DATA_BLOCK "Recipe Libraries"   // DB9
{ S7_Optimized_Access := 'TRUE' }
VERSION : 0.1
   VAR
      me : "Menu: Libraries";
   END_VAR
BEGIN
   me.stations[24].wip[0] := WSTRING#'16.08.208.101.020A$L$$SA DOC Sleeved Before Forming';
   me.stations[24].wip[1] := WSTRING#'16.08.209.031.000C$LDOC Stuffed Shell Before Forming';
   me.stations[24].wip[2] := WSTRING#'16.08.209.091.000D$LSA DPF Stuffed (after Hess)';
   me.stations[24].wip[3] := WSTRING#'16.08.209.233.000E$LSCR Stuffed Shell- NGK Before Forming';
   me.stations[24].wip[4] := WSTRING#'16.08.209.437.000A$LDOC Stuffed Shell Unformed';
   me.stations[24].wip[5] := WSTRING#'16.08.210.031.000B$LStuffed Shell DOC';
   me.stations[24].wip[6] := WSTRING#'16.08.210.421.500A$LStuffed Shell DOC- 2013';
   me.stations[24].wip[7] := WSTRING#'16.08.210.428.000A$LSA DPF Stuffed (after Hess)';
   me.stations[24].wip[8] := WSTRING#'16.08.211.801.400A$L$$SA DOC Sleeved';
   me.stations[24].wip[9] := WSTRING#'16.08.211.801.700B$LDPF Stuffed Shell 1 box longs only';
   me.stations[24].wip[10] := WSTRING#'16.08.211.806.400B$L$$SA DPF Stuffed Shell';
   me.stations[24].wip[11] := WSTRING#'16.08.216.801.600A$LSA DOC Sleeved DDC 2016 unformed';
   me.stations[24].wip[12] := WSTRING#'16.08.216.806.400A$L DPF Sleeved 2016';
   me.stations[24].wip[13] := WSTRING#'16.08.217.408.000A$LSA DPF SLEEVED Hess';
   me.stations[24].wip[14] := WSTRING#'16.08.217.421.500A$LSA DOC SLEEVED - 2HH 2016';
   me.stations[24].wip[15] := WSTRING#'16.08.217.737.000A$LSA DOC SLEEVED - 2V2 2016 unformed';
   me.stations[24].wip[16] := WSTRING#'16.32.307.322.210A$LVolvo - ASSY INLET - SUB 8 Unformed';
   me.stations[24].wip[17] := WSTRING#'16.32.307.332.400A$LAssembly DPF Canning 2016';
   me.stations[24].wip[18] := WSTRING#'16.32.307.472.210A$LSA DOC Canning w/out End Forming';
   me.stations[24].wip[19] := WSTRING#'16.32.407.322.210A$LVOLVO DOC STUFFED SHELL UNFORMED';
   me.stations[24].wip[20] := WSTRING#'16.08.208.081.000H$LDPF Stuffed Shell 1 box longs only';
   me.stations[24].wip[21] := WSTRING#'16.08.208.621.000G$LSA DPF Stuffed Shell';
   me.stations[24].wip[22] := WSTRING#'16.32.407.322.300A$LDPF Stuffed Shell: MD13/MD16';
   me.stations[24].wip[23] := WSTRING#'16.32.307.332.300A$LDPF Stuffed Shell MD11';
   me.stations[25].wip[0] := WSTRING#'16.08.210.421.500A$LStuffed Shell DOC- 2013';
   me.stations[25].wip[1] := WSTRING#'16.08.217.421.500A$LSA DOC SLEEVED - 2HH 2016';
   me.stations[25].wip[2] := WSTRING#'16.08.217.737.000A$LSA DOC SLEEVED - 2V2 2016 unformed';
   me.stations[25].wip[3] := WSTRING#'16.08.208.031.000F$LSCR Stuffed Shell 1 box longs only';
   me.stations[25].wip[4] := WSTRING#'16.08.208.651.000G$LStuffed Shell SCR- NGK';
   me.stations[25].wip[5] := WSTRING#'16.08.211.803.400A$LSCR Stuffed Shell High Power';
   me.stations[25].wip[6] := WSTRING#'16.08.217.233.000A$LSA SCR SLEEVED before FORMING';
   me.stations[25].wip[7] := WSTRING#'16.32.606.411.000A$LStuffed Shell - SCR Horizontal';
   me.stations[25].wip[8] := WSTRING#'16.32.606.421.000A$LStuffed Shell - SCR Horizontal Long- UNI';
   me.stations[25].wip[9] := WSTRING#'16.32.706.311.000A$L$$SCR Stuffed Shell MD11/13: Vert Short';
   me.stations[25].wip[10] := WSTRING#'16.32.706.311.001A$L$$SCR Stuffed Shell MD11/13: Vert Short';
   me.stations[25].wip[11] := WSTRING#'16.32.706.341.000A$LSA SCR Catalyst Module - MD11_MD13 -';
   me.stations[25].wip[12] := WSTRING#'16.32.706.401.000A$LSCR Stuffed Shell MD11/13: Australia';
   me.stations[26].wip[0] := WSTRING#'16.18.015.420.000A$LSA DOC CANNING 11.25 x 5in -END FORMED-';
   me.stations[26].wip[1] := WSTRING#'16.08.211.806.400B$L$$SA DPF Stuffed Shell';
   me.stations[26].wip[2] := WSTRING#'16.08.216.801.600A$LSA DOC Sleeved DDC 2016 unformed';
   me.stations[26].wip[3] := WSTRING#'16.08.216.806.400A$L DPF Sleeved 2016';
   me.stations[26].wip[4] := WSTRING#'16.08.216.751.100A$LSA Sleeved SCR 2016';
   me.stations[26].wip[5] := WSTRING#'16.18.007.300.000A$LSA SCR CANNING 9.5 x 10in -END FORMED-';
   me.stations[26].wip[6] := WSTRING#'16.18.007.310.000A$LSA SCR CANNING 9.5 x 12in -END FORMED-';
   me.stations[26].wip[7] := WSTRING#'16.18.007.320.000B$LSA SCR CANNING 9.5 x 9in -END FORMED-';
   me.stations[26].wip[8] := WSTRING#'16.18.008.300.000A$LSA SCR CANNING 9.5 x 12in -END FORMED-';
   me.stations[26].wip[9] := WSTRING#'16.18.008.310.000A$LSA SCR CANNING 9.5 x 10in -END FORMED-';
   me.stations[26].wip[10] := WSTRING#'16.18.008.320.000A$LSA SCR CANNING 9.5 x 13in -END FORMED-';
   me.stations[26].wip[11] := WSTRING#'16.18.008.340.000A$LSA SCR CANNING 9.5 x 13in -END FORMED-';
   me.stations[26].wip[12] := WSTRING#'16.18.009.301.000H$LSA SCR CANNING 13 x 11in UNFORMED-';
   me.stations[26].wip[13] := WSTRING#'16.18.009.311.000H$LSA SCR CANNING 13 x 12in UNFORMED-';
   me.stations[26].wip[14] := WSTRING#'16.18.009.321.000G$LSA SCR CANNING 13 x 9in UNFORMED';
   me.stations[26].wip[15] := WSTRING#'16.18.009.331.000F$LSA SCR CANNING 13 x 9in UNFORMED';
   me.stations[26].wip[16] := WSTRING#'16.18.009.371.000D$LSA SCR CANNING 13 X10  UNFORMED';
   me.stations[26].wip[17] := WSTRING#'16.18.011.300.000A$LSA SCR CANNING 9.5 x 13.5in -END FORMED-';
   me.stations[26].wip[18] := WSTRING#'16.18.011.310.000A$L SA SCR CANNING 9.5 x 10in -END FORMED-';
   me.stations[26].wip[19] := WSTRING#'16.18.011.320.000A$LSA SCR CANNING 9_5 x 13in -END FORMED-';
   me.stations[26].wip[20] := WSTRING#'16.18.011.330.000A$LSA SCR CANNING 9.5 x 9in -END FORMED-';
   me.stations[26].wip[21] := WSTRING#'16.18.012.400.000A$LSA DOC CANNING 9.5 x 4in -END FORMED_';
   me.stations[26].wip[22] := WSTRING#'16.18.012.410.000A$LSA DOC CANNING 9.5 x 3.3in -END FORMED-';
   me.stations[26].wip[23] := WSTRING#'16.18.012.420.000A$LSA DOC CANNING 9.5 x 4in -END FORMED-';
   me.stations[26].wip[24] := WSTRING#'16.18.012.430.000A$LSA DOC CANNING 9.5 x 3.3in -END FORMED-';
   me.stations[26].wip[25] := WSTRING#'16.18.012.440.000A$LSA DOC CANNING 9.5 x 5in -END FORMED-';
   me.stations[26].wip[26] := WSTRING#'16.18.013.410.000A$LSA DOC CANNING 9_5 x 4_5in -END FORMED-';
   me.stations[26].wip[27] := WSTRING#'16.18.013.420.000A$LSA DOC CANNING 9.5 x 5.5in -END FORMED-';
   me.stations[26].wip[28] := WSTRING#'16.18.015.400.000A$LSA DOC CANNING 11.25 x 4in -END FORMED-';
   me.stations[26].wip[29] := WSTRING#'16.18.015.410.000A$LSA DOC CANNING 11_25 x 5in -END FORMED-';
   me.stations[26].wip[30] := WSTRING#'16.18.015.430.000A$LSA DOC CANNING 11.25 x 3.4in -END FORMED';
   me.stations[26].wip[31] := WSTRING#'16.18.015.450.000A$LSA DOC CANNING 11.25 x 5in -END FORMED-';
   me.stations[26].wip[32] := WSTRING#'16.18.016.400.000A$LSA DOC CANNING 11.25 x 3.4in -END FORMED';
   me.stations[26].wip[33] := WSTRING#'16.18.017.300.000A$LSA SCR CANNING 12 x 10in -END FORMED-';
   me.stations[26].wip[34] := WSTRING#'16.18.017.310.000A$LSA SCR CANNING 12 x 9in -END FORMED-';
   me.stations[26].wip[35] := WSTRING#'16.18.017.321.000F$LSA SCR CANNING 12x7in UNFORMED-';
   me.stations[26].wip[36] := WSTRING#'16.18.018.400.000A$LSA DOC CANNING 11.25 x 6.8in -END FORMED';
   me.stations[26].wip[37] := WSTRING#'16.18.018.410.000A$LSA DOC CANNING 11.25 x 5in -END FORMED-';
   me.stations[26].wip[38] := WSTRING#'16.18.018.420.000A$LSA DOC CANNING 11.25 x 6.8in -END FORMED';
   me.stations[26].wip[39] := WSTRING#'16.18.018.440.000A$LSA DOC CANNING 11.25 x 5in -END FORMED-';
   me.stations[26].wip[40] := WSTRING#'16.18.011.340.000A$LSCR CANNING 9.5 x 9in -END FORMED-';
   me.stations[27].wip[0] := WSTRING#'16.08.211.801.700B$LDPF Stuffed Shell 1 box longs only';
   me.stations[27].wip[1] := WSTRING#'16.32.307.322.210A$LVolvo - ASSY INLET - SUB 8 Unformed';
   me.stations[27].wip[2] := WSTRING#'16.32.606.411.000A$LStuffed Shell - SCR Horizontal';
   me.stations[27].wip[3] := WSTRING#'16.32.112.311.001A$LSA SCR CANNING UNFORMED';
   me.stations[27].wip[4] := WSTRING#'16.32.112.553.300C$LSA SCR CANNING A700 UNFORMED';
   me.stations[27].wip[5] := WSTRING#'16.32.112.304.008A$LASSY SCR CANNING FORMED';
   me.stations[27].wip[6] := WSTRING#'16.32.112.516.000G$LASSY DPF CANNING A700';
   me.stations[27].wip[7] := WSTRING#'16.32.112.543.000E$LASSY DOC CANNING A700';
   me.stations[28].wip[0] := WSTRING#'11.52.001.312.000B$LSA JL 2.2L DPF CANNING';
   me.stations[28].wip[1] := WSTRING#'11.54.007.309.000D$LSTUFFED SHELL ASSEMBLY USA-U625';
   me.stations[28].wip[2] := WSTRING#'11.54.007.309.002D$LSTUFFED SHELL ASSEMBLY USA-U625';
   me.stations[28].wip[3] := WSTRING#'11.54.007.309.009D$LSTUFFED SHELL ASSEMBLY USA-U625';
   me.stations[24].raw[20,7] := WSTRING#'';
   me.stations[24].raw[20,6] := WSTRING#'';
   me.stations[24].raw[20,5] := WSTRING#'';
   me.stations[24].raw[20,4] := WSTRING#'';
   me.stations[24].raw[20,3] := WSTRING#'';
   me.stations[24].raw[20,2] := WSTRING#'16.08.208.091.000A';
   me.stations[24].raw[20,1] := WSTRING#'16.08.208.311.000F';
   me.stations[24].raw[20,0] := WSTRING#'16.08.208.081.010B';
   me.stations[24].raw[19,7] := WSTRING#'';
   me.stations[24].raw[19,6] := WSTRING#'';
   me.stations[24].raw[19,5] := WSTRING#'';
   me.stations[24].raw[19,4] := WSTRING#'';
   me.stations[24].raw[19,3] := WSTRING#'';
   me.stations[24].raw[19,2] := WSTRING#'16.32.407.241.150B';
   me.stations[24].raw[19,1] := WSTRING#'16.32.407.241.170B';
   me.stations[24].raw[19,0] := WSTRING#'16.32.407.441.160A';
   me.stations[24].raw[18,7] := WSTRING#'';
   me.stations[24].raw[18,6] := WSTRING#'';
   me.stations[24].raw[18,5] := WSTRING#'';
   me.stations[24].raw[18,4] := WSTRING#'';
   me.stations[24].raw[18,3] := WSTRING#'';
   me.stations[24].raw[18,2] := WSTRING#'16.32.112.543.020A';
   me.stations[24].raw[18,1] := WSTRING#'16.32.307.211.170B';
   me.stations[24].raw[18,0] := WSTRING#'16.32.307.461.160A';
   me.stations[24].raw[17,7] := WSTRING#'';
   me.stations[24].raw[17,6] := WSTRING#'';
   me.stations[24].raw[17,5] := WSTRING#'';
   me.stations[24].raw[17,4] := WSTRING#'';
   me.stations[24].raw[17,3] := WSTRING#'';
   me.stations[24].raw[17,2] := WSTRING#'16.32.112.536.010A';
   me.stations[24].raw[17,1] := WSTRING#'16.32.307.212.320C';
   me.stations[24].raw[17,0] := WSTRING#'16.32.307.312.310A';
   me.stations[24].raw[16,7] := WSTRING#'';
   me.stations[24].raw[16,6] := WSTRING#'';
   me.stations[24].raw[16,5] := WSTRING#'';
   me.stations[24].raw[16,4] := WSTRING#'';
   me.stations[24].raw[16,3] := WSTRING#'';
   me.stations[24].raw[16,2] := WSTRING#'16.32.307.211.150B';
   me.stations[24].raw[16,1] := WSTRING#'16.32.307.211.170B';
   me.stations[24].raw[16,0] := WSTRING#'16.32.307.461.160A';
   me.stations[24].raw[15,7] := WSTRING#'';
   me.stations[24].raw[15,6] := WSTRING#'';
   me.stations[24].raw[15,5] := WSTRING#'';
   me.stations[24].raw[15,4] := WSTRING#'';
   me.stations[24].raw[15,3] := WSTRING#'';
   me.stations[24].raw[15,2] := WSTRING#'16.08.217.421.130A';
   me.stations[24].raw[15,1] := WSTRING#'16.08.209.031.010C';
   me.stations[24].raw[15,0] := WSTRING#'16.08.209.031.030B';
   me.stations[24].raw[14,7] := WSTRING#'';
   me.stations[24].raw[14,6] := WSTRING#'';
   me.stations[24].raw[14,5] := WSTRING#'';
   me.stations[24].raw[14,4] := WSTRING#'';
   me.stations[24].raw[14,3] := WSTRING#'';
   me.stations[24].raw[14,2] := WSTRING#'16.08.217.421.130A';
   me.stations[24].raw[14,1] := WSTRING#'16.08.210.031.010B';
   me.stations[24].raw[14,0] := WSTRING#'16.08.209.031.030B';
   me.stations[24].raw[13,7] := WSTRING#'';
   me.stations[24].raw[13,6] := WSTRING#'';
   me.stations[24].raw[13,5] := WSTRING#'';
   me.stations[24].raw[13,4] := WSTRING#'';
   me.stations[24].raw[13,3] := WSTRING#'';
   me.stations[24].raw[13,2] := WSTRING#'16.08.217.421.010A';
   me.stations[24].raw[13,1] := WSTRING#'16.08.209.091.010C';
   me.stations[24].raw[13,0] := WSTRING#'16.08.210.421.020A';
   me.stations[24].raw[12,7] := WSTRING#'';
   me.stations[24].raw[12,6] := WSTRING#'';
   me.stations[24].raw[12,5] := WSTRING#'';
   me.stations[24].raw[12,4] := WSTRING#'';
   me.stations[24].raw[12,3] := WSTRING#'';
   me.stations[24].raw[12,2] := WSTRING#'16.08.216.806.020A';
   me.stations[24].raw[12,1] := WSTRING#'16.08.208.631.000F';
   me.stations[24].raw[12,0] := WSTRING#'16.08.216.315.000A';
   me.stations[24].raw[11,7] := WSTRING#'';
   me.stations[24].raw[11,6] := WSTRING#'';
   me.stations[24].raw[11,5] := WSTRING#'';
   me.stations[24].raw[11,4] := WSTRING#'';
   me.stations[24].raw[11,3] := WSTRING#'';
   me.stations[24].raw[11,2] := WSTRING#'16.08.216.053.000A';
   me.stations[24].raw[11,1] := WSTRING#'16.08.208.321.000G';
   me.stations[24].raw[11,0] := WSTRING#'16.08.208.101.010C';
   me.stations[24].raw[10,7] := WSTRING#'';
   me.stations[24].raw[10,6] := WSTRING#'';
   me.stations[24].raw[10,5] := WSTRING#'';
   me.stations[24].raw[10,4] := WSTRING#'';
   me.stations[24].raw[10,3] := WSTRING#'';
   me.stations[24].raw[10,2] := WSTRING#'16.08.211.806.020A';
   me.stations[24].raw[10,1] := WSTRING#'16.08.208.631.000F';
   me.stations[24].raw[10,0] := WSTRING#'16.08.216.315.000A';
   me.stations[24].raw[9,7] := WSTRING#'';
   me.stations[24].raw[9,6] := WSTRING#'';
   me.stations[24].raw[9,5] := WSTRING#'';
   me.stations[24].raw[9,4] := WSTRING#'';
   me.stations[24].raw[9,3] := WSTRING#'';
   me.stations[24].raw[9,2] := WSTRING#'16.08.211.801.020A';
   me.stations[24].raw[9,1] := WSTRING#'16.08.208.631.000F';
   me.stations[24].raw[9,0] := WSTRING#'16.08.216.315.002A';
   me.stations[24].raw[8,7] := WSTRING#'';
   me.stations[24].raw[8,6] := WSTRING#'';
   me.stations[24].raw[8,5] := WSTRING#'';
   me.stations[24].raw[8,4] := WSTRING#'';
   me.stations[24].raw[8,3] := WSTRING#'';
   me.stations[24].raw[8,2] := WSTRING#'16.08.211.801.010A';
   me.stations[24].raw[8,1] := WSTRING#'16.08.208.321.000G';
   me.stations[24].raw[8,0] := WSTRING#'16.08.208.101.010C';
   me.stations[24].raw[7,7] := WSTRING#'';
   me.stations[24].raw[7,6] := WSTRING#'';
   me.stations[24].raw[7,5] := WSTRING#'';
   me.stations[24].raw[7,4] := WSTRING#'';
   me.stations[24].raw[7,3] := WSTRING#'';
   me.stations[24].raw[7,2] := WSTRING#'16.08.210.421.010A';
   me.stations[24].raw[7,1] := WSTRING#'16.08.209.091.010C';
   me.stations[24].raw[7,0] := WSTRING#'16.08.210.421.020A';
   me.stations[24].raw[6,7] := WSTRING#'';
   me.stations[24].raw[6,6] := WSTRING#'';
   me.stations[24].raw[6,5] := WSTRING#'';
   me.stations[24].raw[6,4] := WSTRING#'';
   me.stations[24].raw[6,3] := WSTRING#'';
   me.stations[24].raw[6,2] := WSTRING#'16.08.210.421.030A';
   me.stations[24].raw[6,1] := WSTRING#'16.08.210.031.010B';
   me.stations[24].raw[6,0] := WSTRING#'16.08.209.031.030B';
   me.stations[24].raw[5,7] := WSTRING#'';
   me.stations[24].raw[5,6] := WSTRING#'';
   me.stations[24].raw[5,5] := WSTRING#'';
   me.stations[24].raw[5,4] := WSTRING#'';
   me.stations[24].raw[5,3] := WSTRING#'';
   me.stations[24].raw[5,2] := WSTRING#'16.08.209.031.050A';
   me.stations[24].raw[5,1] := WSTRING#'16.08.210.031.010B';
   me.stations[24].raw[5,0] := WSTRING#'16.08.209.031.030B';
   me.stations[24].raw[4,7] := WSTRING#'';
   me.stations[24].raw[4,6] := WSTRING#'';
   me.stations[24].raw[4,5] := WSTRING#'';
   me.stations[24].raw[4,4] := WSTRING#'';
   me.stations[24].raw[4,3] := WSTRING#'';
   me.stations[24].raw[4,2] := WSTRING#'16.08.210.421.030A';
   me.stations[24].raw[4,1] := WSTRING#'16.08.209.031.010C';
   me.stations[24].raw[4,0] := WSTRING#'16.08.209.031.030B';
   me.stations[24].raw[3,7] := WSTRING#'';
   me.stations[24].raw[3,6] := WSTRING#'';
   me.stations[24].raw[3,5] := WSTRING#'';
   me.stations[24].raw[3,4] := WSTRING#'16.08.208.041.000A';
   me.stations[24].raw[3,3] := WSTRING#'16.08.211.291.000A';
   me.stations[24].raw[3,2] := WSTRING#'16.08.209.232.010C';
   me.stations[24].raw[3,1] := WSTRING#'16.08.208.031.020C';
   me.stations[24].raw[3,0] := WSTRING#'16.08.208.651.010B';
   me.stations[24].raw[2,7] := WSTRING#'';
   me.stations[24].raw[2,6] := WSTRING#'';
   me.stations[24].raw[2,5] := WSTRING#'';
   me.stations[24].raw[2,4] := WSTRING#'';
   me.stations[24].raw[2,3] := WSTRING#'';
   me.stations[24].raw[2,2] := WSTRING#'16.08.209.091.060A';
   me.stations[24].raw[2,1] := WSTRING#'16.08.209.091.010C';
   me.stations[24].raw[2,0] := WSTRING#'16.08.209.091.030D';
   me.stations[24].raw[1,7] := WSTRING#'';
   me.stations[24].raw[1,6] := WSTRING#'';
   me.stations[24].raw[1,5] := WSTRING#'';
   me.stations[24].raw[1,4] := WSTRING#'';
   me.stations[24].raw[1,3] := WSTRING#'';
   me.stations[24].raw[1,2] := WSTRING#'16.08.209.031.050A';
   me.stations[24].raw[1,1] := WSTRING#'16.08.209.031.010C';
   me.stations[24].raw[1,0] := WSTRING#'16.08.209.031.030B';
   me.stations[24].raw[0,7] := WSTRING#'';
   me.stations[24].raw[0,6] := WSTRING#'';
   me.stations[24].raw[0,5] := WSTRING#'';
   me.stations[24].raw[0,4] := WSTRING#'';
   me.stations[24].raw[0,3] := WSTRING#'';
   me.stations[24].raw[0,2] := WSTRING#'16.08.208.111.000B';
   me.stations[24].raw[0,1] := WSTRING#'16.08.208.321.000G';
   me.stations[24].raw[0,0] := WSTRING#'16.08.208.101.010C';
   me.stations[26].raw[15,6] := WSTRING#'';
   me.stations[26].raw[15,5] := WSTRING#'';
   me.stations[26].raw[15,4] := WSTRING#'16.18.009.331.050A';
   me.stations[26].raw[15,3] := WSTRING#'16.18.009.321.030A';
   me.stations[26].raw[15,2] := WSTRING#'16.18.009.321.010A';
   me.stations[26].raw[15,1] := WSTRING#'16.18.009.321.020B';
   me.stations[26].raw[15,0] := WSTRING#'16.18.009.301.020B';
   me.stations[26].raw[14,7] := WSTRING#'';
   me.stations[26].raw[14,6] := WSTRING#'';
   me.stations[26].raw[14,5] := WSTRING#'';
   me.stations[26].raw[14,4] := WSTRING#'16.18.009.321.030A';
   me.stations[26].raw[14,3] := WSTRING#'16.18.009.321.010A';
   me.stations[26].raw[14,2] := WSTRING#'16.18.009.301.050A';
   me.stations[26].raw[14,1] := WSTRING#'16.18.009.301.020B';
   me.stations[26].raw[14,0] := WSTRING#'16.18.009.321.020B';
   me.stations[26].raw[13,7] := WSTRING#'';
   me.stations[26].raw[13,6] := WSTRING#'';
   me.stations[26].raw[13,5] := WSTRING#'';
   me.stations[26].raw[13,4] := WSTRING#'';
   me.stations[26].raw[13,3] := WSTRING#'16.18.009.301.030A';
   me.stations[26].raw[13,2] := WSTRING#'16.18.009.311.010A';
   me.stations[26].raw[13,1] := WSTRING#'16.18.009.301.050A';
   me.stations[26].raw[13,0] := WSTRING#'16.18.009.301.040B';
   me.stations[26].raw[12,7] := WSTRING#'';
   me.stations[26].raw[12,6] := WSTRING#'';
   me.stations[26].raw[12,5] := WSTRING#'';
   me.stations[26].raw[12,4] := WSTRING#'16.18.009.301.030A';
   me.stations[26].raw[12,3] := WSTRING#'16.18.009.301.010A';
   me.stations[26].raw[12,2] := WSTRING#'16.18.009.301.050A';
   me.stations[26].raw[12,1] := WSTRING#'16.18.009.301.040B';
   me.stations[26].raw[12,0] := WSTRING#'16.18.009.301.020B';
   me.stations[26].raw[11,7] := WSTRING#'';
   me.stations[26].raw[11,6] := WSTRING#'';
   me.stations[26].raw[11,5] := WSTRING#'';
   me.stations[26].raw[11,4] := WSTRING#'';
   me.stations[26].raw[11,3] := WSTRING#'';
   me.stations[26].raw[11,2] := WSTRING#'16.18.008.311.010A';
   me.stations[26].raw[11,1] := WSTRING#'16.18.008.301.030A';
   me.stations[26].raw[11,0] := WSTRING#'16.18.008.311.020B';
   me.stations[26].raw[10,7] := WSTRING#'';
   me.stations[26].raw[10,6] := WSTRING#'';
   me.stations[26].raw[10,5] := WSTRING#'';
   me.stations[26].raw[10,4] := WSTRING#'16.18.008.301.020A';
   me.stations[26].raw[10,3] := WSTRING#'16.18.007.301.010A';
   me.stations[26].raw[10,2] := WSTRING#'16.18.008.301.030A';
   me.stations[26].raw[10,1] := WSTRING#'16.18.011.321.020B';
   me.stations[26].raw[10,0] := WSTRING#'16.18.011.301.020B';
   me.stations[26].raw[9,7] := WSTRING#'';
   me.stations[26].raw[9,6] := WSTRING#'';
   me.stations[26].raw[9,5] := WSTRING#'';
   me.stations[26].raw[9,4] := WSTRING#'';
   me.stations[26].raw[9,3] := WSTRING#'16.18.011.321.010A';
   me.stations[26].raw[9,2] := WSTRING#'16.18.007.301.010A';
   me.stations[26].raw[9,1] := WSTRING#'16.18.008.301.030A';
   me.stations[26].raw[9,0] := WSTRING#'16.18.011.321.020B';
   me.stations[26].raw[8,7] := WSTRING#'';
   me.stations[26].raw[8,6] := WSTRING#'';
   me.stations[26].raw[8,5] := WSTRING#'';
   me.stations[26].raw[8,4] := WSTRING#'16.18.008.301.020A';
   me.stations[26].raw[8,3] := WSTRING#'16.18.008.301.010A';
   me.stations[26].raw[8,2] := WSTRING#'16.18.008.301.030A';
   me.stations[26].raw[8,1] := WSTRING#'16.18.011.301.020B';
   me.stations[26].raw[8,0] := WSTRING#'16.18.012.401.020A';
   me.stations[26].raw[7,7] := WSTRING#'';
   me.stations[26].raw[7,6] := WSTRING#'';
   me.stations[26].raw[7,5] := WSTRING#'';
   me.stations[26].raw[7,4] := WSTRING#'16.18.007.311.010A';
   me.stations[26].raw[7,3] := WSTRING#'16.18.007.301.010A';
   me.stations[26].raw[7,2] := WSTRING#'16.18.007.321.010B';
   me.stations[26].raw[7,1] := WSTRING#'16.18.011.321.020B';
   me.stations[26].raw[7,0] := WSTRING#'16.18.012.401.020A';
   me.stations[26].raw[6,7] := WSTRING#'';
   me.stations[26].raw[6,6] := WSTRING#'';
   me.stations[26].raw[6,5] := WSTRING#'';
   me.stations[26].raw[6,4] := WSTRING#'16.18.007.311.010A';
   me.stations[26].raw[6,3] := WSTRING#'16.18.011.301.010A';
   me.stations[26].raw[6,2] := WSTRING#'16.18.007.311.020A';
   me.stations[26].raw[6,1] := WSTRING#'16.18.011.301.020B';
   me.stations[26].raw[6,0] := WSTRING#'16.18.012.401.020A';
   me.stations[26].raw[5,7] := WSTRING#'';
   me.stations[26].raw[5,6] := WSTRING#'';
   me.stations[26].raw[5,5] := WSTRING#'';
   me.stations[26].raw[5,4] := WSTRING#'';
   me.stations[26].raw[5,3] := WSTRING#'16.18.007.301.010A';
   me.stations[26].raw[5,2] := WSTRING#'16.18.011.321.010A';
   me.stations[26].raw[5,1] := WSTRING#'16.18.007.301.020A';
   me.stations[26].raw[5,0] := WSTRING#'16.18.011.321.020B';
   me.stations[26].raw[4,7] := WSTRING#'';
   me.stations[26].raw[4,6] := WSTRING#'';
   me.stations[26].raw[4,5] := WSTRING#'';
   me.stations[26].raw[4,4] := WSTRING#'16.08.216.057.001A';
   me.stations[26].raw[4,3] := WSTRING#'16.08.216.291.000A';
   me.stations[26].raw[4,2] := WSTRING#'16.08.208.661.000F';
   me.stations[26].raw[4,1] := WSTRING#'16.08.216.315.001A';
   me.stations[26].raw[4,0] := WSTRING#'16.08.216.315.002A';
   me.stations[26].raw[3,7] := WSTRING#'';
   me.stations[26].raw[3,6] := WSTRING#'';
   me.stations[26].raw[3,5] := WSTRING#'';
   me.stations[26].raw[3,4] := WSTRING#'';
   me.stations[26].raw[3,3] := WSTRING#'';
   me.stations[26].raw[3,2] := WSTRING#'16.08.216.806.020A';
   me.stations[26].raw[3,1] := WSTRING#'16.08.208.631.000F';
   me.stations[26].raw[3,0] := WSTRING#'16.08.216.315.000A';
   me.stations[26].raw[2,7] := WSTRING#'';
   me.stations[26].raw[2,6] := WSTRING#'';
   me.stations[26].raw[2,5] := WSTRING#'';
   me.stations[26].raw[2,4] := WSTRING#'';
   me.stations[26].raw[2,3] := WSTRING#'';
   me.stations[26].raw[2,2] := WSTRING#'16.08.216.053.000A';
   me.stations[26].raw[2,1] := WSTRING#'16.08.208.321.000G';
   me.stations[26].raw[2,0] := WSTRING#'16.08.208.101.010C';
   me.stations[26].raw[1,7] := WSTRING#'';
   me.stations[26].raw[1,6] := WSTRING#'';
   me.stations[26].raw[1,5] := WSTRING#'';
   me.stations[26].raw[1,4] := WSTRING#'';
   me.stations[26].raw[1,3] := WSTRING#'';
   me.stations[26].raw[1,2] := WSTRING#'16.08.211.806.020A';
   me.stations[26].raw[1,1] := WSTRING#'16.08.208.631.000F';
   me.stations[26].raw[1,0] := WSTRING#'16.08.216.315.000A';
   me.stations[26].raw[0,7] := WSTRING#'';
   me.stations[26].raw[0,6] := WSTRING#'';
   me.stations[26].raw[0,5] := WSTRING#'';
   me.stations[26].raw[0,4] := WSTRING#'';
   me.stations[26].raw[0,3] := WSTRING#'';
   me.stations[26].raw[0,2] := WSTRING#'16.18.015.421.010A';
   me.stations[26].raw[0,1] := WSTRING#'16.18.015.411.030A';
   me.stations[26].raw[0,0] := WSTRING#'16.18.015.421.020B';
   me.stations[24].raw[23,7] := WSTRING#'';
   me.stations[24].raw[23,6] := WSTRING#'';
   me.stations[24].raw[23,5] := WSTRING#'';
   me.stations[24].raw[23,4] := WSTRING#'';
   me.stations[24].raw[23,3] := WSTRING#'';
   me.stations[24].raw[23,2] := WSTRING#'16.32.307.232.300B';
   me.stations[24].raw[23,1] := WSTRING#'16.32.307.212.320C';
   me.stations[24].raw[23,0] := WSTRING#'16.32.307.312.310A';
   me.stations[24].raw[22,7] := WSTRING#'';
   me.stations[24].raw[22,6] := WSTRING#'';
   me.stations[24].raw[22,5] := WSTRING#'';
   me.stations[24].raw[22,4] := WSTRING#'';
   me.stations[24].raw[22,3] := WSTRING#'';
   me.stations[24].raw[22,2] := WSTRING#'16.32.307.262.300B';
   me.stations[24].raw[22,1] := WSTRING#'16.32.307.212.320C';
   me.stations[24].raw[22,0] := WSTRING#'16.32.307.312.310A';
   me.stations[24].raw[21,7] := WSTRING#'';
   me.stations[24].raw[21,6] := WSTRING#'';
   me.stations[24].raw[21,5] := WSTRING#'';
   me.stations[24].raw[21,4] := WSTRING#'';
   me.stations[24].raw[21,3] := WSTRING#'';
   me.stations[24].raw[21,2] := WSTRING#'16.08.211.781.000A';
   me.stations[24].raw[21,1] := WSTRING#'16.08.208.631.000F';
   me.stations[24].raw[21,0] := WSTRING#'16.08.208.621.010C';
   me.stations[25].raw[12,7] := WSTRING#'';
   me.stations[25].raw[12,6] := WSTRING#'';
   me.stations[25].raw[12,5] := WSTRING#'';
   me.stations[25].raw[12,4] := WSTRING#'';
   me.stations[25].raw[12,3] := WSTRING#'16.32.706.401.050A';
   me.stations[25].raw[12,2] := WSTRING#'16.32.706.401.040A';
   me.stations[25].raw[12,1] := WSTRING#'16.32.706.321.010B';
   me.stations[25].raw[12,0] := WSTRING#'16.32.706.321.030B';
   me.stations[25].raw[11,7] := WSTRING#'';
   me.stations[25].raw[11,6] := WSTRING#'';
   me.stations[25].raw[11,5] := WSTRING#'';
   me.stations[25].raw[11,4] := WSTRING#'';
   me.stations[25].raw[11,3] := WSTRING#'16.32.112.553.010A';
   me.stations[25].raw[11,2] := WSTRING#'16.32.112.553.020A';
   me.stations[25].raw[11,1] := WSTRING#'16.32.706.311.010C';
   me.stations[25].raw[11,0] := WSTRING#'16.32.706.311.020B';
   me.stations[25].raw[10,7] := WSTRING#'';
   me.stations[25].raw[10,6] := WSTRING#'';
   me.stations[25].raw[10,5] := WSTRING#'';
   me.stations[25].raw[10,4] := WSTRING#'';
   me.stations[25].raw[10,3] := WSTRING#'16.32.112.057.010A';
   me.stations[25].raw[10,2] := WSTRING#'16.32.112.054.041A';
   me.stations[25].raw[10,1] := WSTRING#'16.32.706.311.010C';
   me.stations[25].raw[10,0] := WSTRING#'16.32.706.311.020B';
   me.stations[25].raw[9,7] := WSTRING#'';
   me.stations[25].raw[9,6] := WSTRING#'';
   me.stations[25].raw[9,5] := WSTRING#'';
   me.stations[25].raw[9,4] := WSTRING#'';
   me.stations[25].raw[9,3] := WSTRING#'16.32.706.311.050B';
   me.stations[25].raw[9,2] := WSTRING#'16.32.706.311.040B';
   me.stations[25].raw[9,1] := WSTRING#'16.32.706.311.010C';
   me.stations[25].raw[9,0] := WSTRING#'16.32.706.311.020B';
   me.stations[25].raw[8,7] := WSTRING#'';
   me.stations[25].raw[8,6] := WSTRING#'';
   me.stations[25].raw[8,5] := WSTRING#'';
   me.stations[25].raw[8,4] := WSTRING#'';
   me.stations[25].raw[8,3] := WSTRING#'16.32.606.311.050B';
   me.stations[25].raw[8,2] := WSTRING#'16.32.606.321.030B';
   me.stations[25].raw[8,1] := WSTRING#'16.32.606.321.010B';
   me.stations[25].raw[8,0] := WSTRING#'16.32.606.311.070A';
   me.stations[25].raw[7,7] := WSTRING#'';
   me.stations[25].raw[7,6] := WSTRING#'';
   me.stations[25].raw[7,5] := WSTRING#'';
   me.stations[25].raw[7,4] := WSTRING#'16.32.606.311.050B';
   me.stations[25].raw[7,3] := WSTRING#'16.32.606.311.040B';
   me.stations[25].raw[7,2] := WSTRING#'16.32.606.311.010C';
   me.stations[25].raw[7,1] := WSTRING#'16.32.606.311.070A';
   me.stations[25].raw[7,0] := WSTRING#'16.32.606.311.060A';
   me.stations[25].raw[6,7] := WSTRING#'';
   me.stations[25].raw[6,6] := WSTRING#'';
   me.stations[25].raw[6,5] := WSTRING#'';
   me.stations[25].raw[6,4] := WSTRING#'16.08.216.057.001A';
   me.stations[25].raw[6,3] := WSTRING#'16.08.216.291.000A';
   me.stations[25].raw[6,2] := WSTRING#'16.08.209.232.010C';
   me.stations[25].raw[6,1] := WSTRING#'16.08.216.315.002A';
   me.stations[25].raw[6,0] := WSTRING#'16.08.216.315.001A';
   me.stations[25].raw[5,7] := WSTRING#'';
   me.stations[25].raw[5,6] := WSTRING#'';
   me.stations[25].raw[5,5] := WSTRING#'';
   me.stations[25].raw[5,4] := WSTRING#'';
   me.stations[25].raw[5,3] := WSTRING#'16.08.208.051.000A';
   me.stations[25].raw[5,2] := WSTRING#'16.08.208.041.000A';
   me.stations[25].raw[5,1] := WSTRING#'16.08.208.661.000F';
   me.stations[25].raw[5,0] := WSTRING#'16.08.208.031.020C';
   me.stations[25].raw[4,7] := WSTRING#'';
   me.stations[25].raw[4,6] := WSTRING#'';
   me.stations[25].raw[4,5] := WSTRING#'';
   me.stations[25].raw[4,4] := WSTRING#'16.08.211.291.000A';
   me.stations[25].raw[4,3] := WSTRING#'16.08.208.041.000A';
   me.stations[25].raw[4,2] := WSTRING#'16.08.208.661.000F';
   me.stations[25].raw[4,1] := WSTRING#'16.08.208.031.020C';
   me.stations[25].raw[4,0] := WSTRING#'16.08.208.651.010B';
   me.stations[25].raw[3,7] := WSTRING#'';
   me.stations[25].raw[3,6] := WSTRING#'';
   me.stations[25].raw[3,5] := WSTRING#'';
   me.stations[25].raw[3,4] := WSTRING#'';
   me.stations[25].raw[3,3] := WSTRING#'16.08.208.051.000A';
   me.stations[25].raw[3,2] := WSTRING#'16.08.208.041.000A';
   me.stations[25].raw[3,1] := WSTRING#'16.08.208.301.000F';
   me.stations[25].raw[3,0] := WSTRING#'16.08.208.031.020C';
   me.stations[25].raw[2,7] := WSTRING#'';
   me.stations[25].raw[2,6] := WSTRING#'';
   me.stations[25].raw[2,5] := WSTRING#'';
   me.stations[25].raw[2,4] := WSTRING#'';
   me.stations[25].raw[2,3] := WSTRING#'';
   me.stations[25].raw[2,2] := WSTRING#'16.08.217.421.130A';
   me.stations[25].raw[2,1] := WSTRING#'16.08.209.031.010C';
   me.stations[25].raw[2,0] := WSTRING#'16.08.209.031.030B';
   me.stations[25].raw[1,7] := WSTRING#'';
   me.stations[25].raw[1,6] := WSTRING#'';
   me.stations[25].raw[1,5] := WSTRING#'';
   me.stations[25].raw[1,4] := WSTRING#'';
   me.stations[25].raw[1,3] := WSTRING#'';
   me.stations[25].raw[1,2] := WSTRING#'16.08.217.421.130A';
   me.stations[25].raw[1,1] := WSTRING#'16.08.210.031.010B';
   me.stations[25].raw[1,0] := WSTRING#'16.08.209.031.030B';
   me.stations[25].raw[0,7] := WSTRING#'';
   me.stations[25].raw[0,6] := WSTRING#'';
   me.stations[25].raw[0,5] := WSTRING#'';
   me.stations[25].raw[0,4] := WSTRING#'';
   me.stations[25].raw[0,3] := WSTRING#'';
   me.stations[25].raw[0,2] := WSTRING#'16.08.210.421.030A';
   me.stations[25].raw[0,1] := WSTRING#'16.08.210.031.010B';
   me.stations[25].raw[0,0] := WSTRING#'16.08.209.031.030B';
   me.stations[26].raw[15,7] := WSTRING#'';
   me.stations[26].raw[16,0] := WSTRING#'16.18.009.301.020B';
   me.stations[26].raw[16,1] := WSTRING#'16.18.009.301.050A';
   me.stations[26].raw[16,2] := WSTRING#'16.18.009.331.030A';
   me.stations[26].raw[16,3] := WSTRING#'16.18.009.371.010A';
   me.stations[26].raw[16,4] := WSTRING#'';
   me.stations[26].raw[16,5] := WSTRING#'';
   me.stations[26].raw[16,6] := WSTRING#'';
   me.stations[26].raw[16,7] := WSTRING#'';
   me.stations[26].raw[17,0] := WSTRING#'16.18.011.301.020B';
   me.stations[26].raw[17,1] := WSTRING#'16.18.011.301.040B';
   me.stations[26].raw[17,2] := WSTRING#'16.18.008.301.030A';
   me.stations[26].raw[17,3] := WSTRING#'16.18.011.301.030A';
   me.stations[26].raw[17,4] := WSTRING#'16.18.011.301.010A';
   me.stations[26].raw[17,5] := WSTRING#'';
   me.stations[26].raw[17,6] := WSTRING#'';
   me.stations[26].raw[17,7] := WSTRING#'';
   me.stations[26].raw[18,0] := WSTRING#'16.18.011.321.020B';
   me.stations[26].raw[18,1] := WSTRING#'16.18.011.311.020A';
   me.stations[26].raw[18,2] := WSTRING#'16.18.007.301.010A';
   me.stations[26].raw[18,3] := WSTRING#'16.18.011.321.010A';
   me.stations[26].raw[18,4] := WSTRING#'';
   me.stations[26].raw[18,5] := WSTRING#'';
   me.stations[26].raw[18,6] := WSTRING#'';
   me.stations[26].raw[18,7] := WSTRING#'';
   me.stations[26].raw[19,0] := WSTRING#'16.18.011.321.020B';
   me.stations[26].raw[19,1] := WSTRING#'16.18.011.301.020B';
   me.stations[26].raw[19,2] := WSTRING#'16.18.011.321.030A';
   me.stations[26].raw[19,3] := WSTRING#'16.18.011.321.010A';
   me.stations[26].raw[19,4] := WSTRING#'16.18.011.301.010A';
   me.stations[26].raw[19,5] := WSTRING#'';
   me.stations[26].raw[19,6] := WSTRING#'';
   me.stations[26].raw[19,7] := WSTRING#'';
   me.stations[26].raw[20,0] := WSTRING#'16.18.011.331.020D';
   me.stations[26].raw[20,1] := WSTRING#'16.18.011.311.020A';
   me.stations[26].raw[20,2] := WSTRING#'16.18.011.331.010A';
   me.stations[26].raw[20,3] := WSTRING#'';
   me.stations[26].raw[20,4] := WSTRING#'';
   me.stations[26].raw[20,5] := WSTRING#'';
   me.stations[26].raw[20,6] := WSTRING#'';
   me.stations[26].raw[20,7] := WSTRING#'';
   me.stations[26].raw[21,0] := WSTRING#'16.18.012.401.020A';
   me.stations[26].raw[21,1] := WSTRING#'16.18.014.411.030A';
   me.stations[26].raw[21,2] := WSTRING#'16.18.012.401.010A';
   me.stations[26].raw[21,3] := WSTRING#'';
   me.stations[26].raw[21,4] := WSTRING#'';
   me.stations[26].raw[21,5] := WSTRING#'';
   me.stations[26].raw[21,6] := WSTRING#'';
   me.stations[26].raw[21,7] := WSTRING#'';
   me.stations[26].raw[22,0] := WSTRING#'16.18.012.411.020B';
   me.stations[26].raw[22,1] := WSTRING#'16.18.014.411.030A';
   me.stations[26].raw[22,2] := WSTRING#'16.18.012.411.010A';
   me.stations[26].raw[22,3] := WSTRING#'';
   me.stations[26].raw[22,4] := WSTRING#'';
   me.stations[26].raw[22,5] := WSTRING#'';
   me.stations[26].raw[22,6] := WSTRING#'';
   me.stations[26].raw[22,7] := WSTRING#'';
   me.stations[26].raw[23,0] := WSTRING#'16.18.012.401.020A';
   me.stations[26].raw[23,1] := WSTRING#'16.18.014.411.030A';
   me.stations[26].raw[23,2] := WSTRING#'16.18.014.411.010A';
   me.stations[26].raw[23,3] := WSTRING#'';
   me.stations[26].raw[23,4] := WSTRING#'';
   me.stations[26].raw[23,5] := WSTRING#'';
   me.stations[26].raw[23,6] := WSTRING#'';
   me.stations[26].raw[23,7] := WSTRING#'';
   me.stations[26].raw[24,0] := WSTRING#'16.18.012.411.020B';
   me.stations[26].raw[24,1] := WSTRING#'16.18.014.411.030A';
   me.stations[26].raw[24,2] := WSTRING#'16.18.012.431.010A';
   me.stations[26].raw[24,3] := WSTRING#'';
   me.stations[26].raw[24,4] := WSTRING#'';
   me.stations[26].raw[24,5] := WSTRING#'';
   me.stations[26].raw[24,6] := WSTRING#'';
   me.stations[26].raw[24,7] := WSTRING#'';
   me.stations[26].raw[25,0] := WSTRING#'16.18.011.321.020B';
   me.stations[26].raw[25,1] := WSTRING#'16.18.013.411.030A';
   me.stations[26].raw[25,2] := WSTRING#'16.18.012.441.010A';
   me.stations[26].raw[25,3] := WSTRING#'';
   me.stations[26].raw[25,4] := WSTRING#'';
   me.stations[26].raw[25,5] := WSTRING#'';
   me.stations[26].raw[25,6] := WSTRING#'';
   me.stations[26].raw[25,7] := WSTRING#'';
   me.stations[26].raw[26,0] := WSTRING#'16.18.013.411.030A';
   me.stations[26].raw[26,1] := WSTRING#'16.18.013.411.010A';
   me.stations[26].raw[26,2] := WSTRING#'16.18.013.411.020B';
   me.stations[26].raw[26,3] := WSTRING#'';
   me.stations[26].raw[26,4] := WSTRING#'';
   me.stations[26].raw[26,5] := WSTRING#'';
   me.stations[26].raw[26,6] := WSTRING#'';
   me.stations[26].raw[26,7] := WSTRING#'';
   me.stations[26].raw[27,0] := WSTRING#'16.18.011.301.040B';
   me.stations[26].raw[27,1] := WSTRING#'16.18.013.411.030A';
   me.stations[26].raw[27,2] := WSTRING#'16.18.013.421.010A';
   me.stations[26].raw[27,3] := WSTRING#'';
   me.stations[26].raw[27,4] := WSTRING#'';
   me.stations[26].raw[27,5] := WSTRING#'';
   me.stations[26].raw[27,6] := WSTRING#'';
   me.stations[26].raw[27,7] := WSTRING#'';
   me.stations[26].raw[28,0] := WSTRING#'16.18.015.421.020B';
   me.stations[26].raw[28,1] := WSTRING#'16.18.015.401.010A';
   me.stations[26].raw[28,2] := WSTRING#'16.18.015.421.010A';
   me.stations[26].raw[28,3] := WSTRING#'';
   me.stations[26].raw[28,4] := WSTRING#'';
   me.stations[26].raw[28,5] := WSTRING#'';
   me.stations[26].raw[28,6] := WSTRING#'';
   me.stations[26].raw[28,7] := WSTRING#'';
   me.stations[26].raw[29,0] := WSTRING#'16.18.015.411.020B';
   me.stations[26].raw[29,1] := WSTRING#'16.18.015.411.030A';
   me.stations[26].raw[29,2] := WSTRING#'16.18.015.411.010A';
   me.stations[26].raw[29,3] := WSTRING#'';
   me.stations[26].raw[29,4] := WSTRING#'';
   me.stations[26].raw[29,5] := WSTRING#'';
   me.stations[26].raw[29,6] := WSTRING#'';
   me.stations[26].raw[29,7] := WSTRING#'';
   me.stations[26].raw[30,0] := WSTRING#'16.18.018.401.020B';
   me.stations[26].raw[30,1] := WSTRING#'16.18.015.401.010A';
   me.stations[26].raw[30,2] := WSTRING#'16.18.018.401.010A';
   me.stations[26].raw[30,3] := WSTRING#'';
   me.stations[26].raw[30,4] := WSTRING#'';
   me.stations[26].raw[30,5] := WSTRING#'';
   me.stations[26].raw[30,6] := WSTRING#'';
   me.stations[26].raw[30,7] := WSTRING#'';
   me.stations[26].raw[31,0] := WSTRING#'16.18.015.411.020B';
   me.stations[26].raw[31,1] := WSTRING#'16.18.015.411.030A';
   me.stations[26].raw[31,2] := WSTRING#'16.18.018.421.010B';
   me.stations[26].raw[31,3] := WSTRING#'';
   me.stations[26].raw[31,4] := WSTRING#'';
   me.stations[26].raw[31,5] := WSTRING#'';
   me.stations[26].raw[31,6] := WSTRING#'';
   me.stations[26].raw[31,7] := WSTRING#'';
   me.stations[26].raw[32,0] := WSTRING#'16.18.018.401.020B';
   me.stations[26].raw[32,1] := WSTRING#'16.18.015.411.030A';
   me.stations[26].raw[32,2] := WSTRING#'16.18.018.401.010A';
   me.stations[26].raw[32,3] := WSTRING#'';
   me.stations[26].raw[32,4] := WSTRING#'';
   me.stations[26].raw[32,5] := WSTRING#'';
   me.stations[26].raw[32,6] := WSTRING#'';
   me.stations[26].raw[32,7] := WSTRING#'';
   me.stations[26].raw[33,0] := WSTRING#'16.18.017.301.040A';
   me.stations[26].raw[33,1] := WSTRING#'16.18.017.301.020A';
   me.stations[26].raw[33,2] := WSTRING#'16.18.017.301.050A';
   me.stations[26].raw[33,3] := WSTRING#'16.18.017.301.030A';
   me.stations[26].raw[33,4] := WSTRING#'16.18.017.301.010A';
   me.stations[26].raw[33,5] := WSTRING#'';
   me.stations[26].raw[33,6] := WSTRING#'';
   me.stations[26].raw[33,7] := WSTRING#'';
   me.stations[26].raw[34,0] := WSTRING#'16.18.017.301.040A';
   me.stations[26].raw[34,1] := WSTRING#'16.18.017.301.050A';
   me.stations[26].raw[34,2] := WSTRING#'16.18.017.301.030A';
   me.stations[26].raw[34,3] := WSTRING#'16.18.017.311.010A';
   me.stations[26].raw[34,4] := WSTRING#'';
   me.stations[26].raw[34,5] := WSTRING#'';
   me.stations[26].raw[34,6] := WSTRING#'';
   me.stations[26].raw[34,7] := WSTRING#'';
   me.stations[26].raw[35,0] := WSTRING#'16.18.017.321.020A';
   me.stations[26].raw[35,1] := WSTRING#'16.18.017.301.050A';
   me.stations[26].raw[35,2] := WSTRING#'16.18.017.321.010A';
   me.stations[26].raw[35,3] := WSTRING#'';
   me.stations[26].raw[35,4] := WSTRING#'';
   me.stations[26].raw[35,5] := WSTRING#'';
   me.stations[26].raw[35,6] := WSTRING#'';
   me.stations[26].raw[35,7] := WSTRING#'';
   me.stations[26].raw[36,0] := WSTRING#'16.18.018.401.020B';
   me.stations[26].raw[36,1] := WSTRING#'16.18.018.401.030A';
   me.stations[26].raw[36,2] := WSTRING#'16.18.018.401.010A';
   me.stations[26].raw[36,3] := WSTRING#'';
   me.stations[26].raw[36,4] := WSTRING#'';
   me.stations[26].raw[36,5] := WSTRING#'';
   me.stations[26].raw[36,6] := WSTRING#'';
   me.stations[26].raw[36,7] := WSTRING#'';
   me.stations[26].raw[37,0] := WSTRING#'16.18.018.401.020B';
   me.stations[26].raw[37,1] := WSTRING#'16.18.018.401.030A';
   me.stations[26].raw[37,2] := WSTRING#'16.18.018.400.000A';
   me.stations[26].raw[37,3] := WSTRING#'';
   me.stations[26].raw[37,4] := WSTRING#'';
   me.stations[26].raw[37,5] := WSTRING#'';
   me.stations[26].raw[37,6] := WSTRING#'';
   me.stations[26].raw[37,7] := WSTRING#'';
   me.stations[26].raw[38,0] := WSTRING#'16.18.018.401.020B';
   me.stations[26].raw[38,1] := WSTRING#'16.18.018.401.030A';
   me.stations[26].raw[38,2] := WSTRING#'16.18.018.411.010A';
   me.stations[26].raw[38,3] := WSTRING#'';
   me.stations[26].raw[38,4] := WSTRING#'';
   me.stations[26].raw[38,5] := WSTRING#'';
   me.stations[26].raw[38,6] := WSTRING#'';
   me.stations[26].raw[38,7] := WSTRING#'';
   me.stations[26].raw[39,0] := WSTRING#'16.18.015.411.020B';
   me.stations[26].raw[39,1] := WSTRING#'16.18.018.401.030A';
   me.stations[26].raw[39,2] := WSTRING#'16.18.018.421.010B';
   me.stations[26].raw[39,3] := WSTRING#'';
   me.stations[26].raw[39,4] := WSTRING#'';
   me.stations[26].raw[39,5] := WSTRING#'';
   me.stations[26].raw[39,6] := WSTRING#'';
   me.stations[26].raw[39,7] := WSTRING#'';
   me.stations[26].raw[40,0] := WSTRING#'16.18.012.401.020A';
   me.stations[26].raw[40,1] := WSTRING#'16.18.011.321.020B';
   me.stations[26].raw[40,2] := WSTRING#'16.18.011.311.020A';
   me.stations[26].raw[40,3] := WSTRING#'16.18.008.301.010A';
   me.stations[26].raw[40,4] := WSTRING#'16.18.011.321.010A';
   me.stations[26].raw[40,5] := WSTRING#'';
   me.stations[26].raw[40,6] := WSTRING#'';
   me.stations[26].raw[40,7] := WSTRING#'';
   me.stations[27].raw[0,0] := WSTRING#'16.08.216.315.002A';
   me.stations[27].raw[0,1] := WSTRING#'16.08.208.631.000F';
   me.stations[27].raw[0,2] := WSTRING#'16.08.211.801.020A';
   me.stations[27].raw[0,3] := WSTRING#'';
   me.stations[27].raw[0,4] := WSTRING#'';
   me.stations[27].raw[0,5] := WSTRING#'';
   me.stations[27].raw[0,6] := WSTRING#'';
   me.stations[27].raw[0,7] := WSTRING#'';
   me.stations[27].raw[1,0] := WSTRING#'16.32.307.461.160A';
   me.stations[27].raw[1,1] := WSTRING#'16.32.307.211.170B';
   me.stations[27].raw[1,2] := WSTRING#'16.32.307.211.150B';
   me.stations[27].raw[1,3] := WSTRING#'';
   me.stations[27].raw[1,4] := WSTRING#'';
   me.stations[27].raw[1,5] := WSTRING#'';
   me.stations[27].raw[1,6] := WSTRING#'';
   me.stations[27].raw[1,7] := WSTRING#'';
   me.stations[27].raw[2,0] := WSTRING#'16.32.606.311.060A';
   me.stations[27].raw[2,1] := WSTRING#'16.32.606.311.070A';
   me.stations[27].raw[2,2] := WSTRING#'16.32.606.311.010C';
   me.stations[27].raw[2,3] := WSTRING#'16.32.606.311.040B';
   me.stations[27].raw[2,4] := WSTRING#'16.32.606.311.050B';
   me.stations[27].raw[2,5] := WSTRING#'';
   me.stations[27].raw[2,6] := WSTRING#'';
   me.stations[27].raw[2,7] := WSTRING#'';
   me.stations[27].raw[3,0] := WSTRING#'16.32.112.553.220A';
   me.stations[27].raw[3,1] := WSTRING#'16.32.112.553.100D';
   me.stations[27].raw[3,2] := WSTRING#'16.32.112.054.041A';
   me.stations[27].raw[3,3] := WSTRING#'16.32.112.057.010A';
   me.stations[27].raw[3,4] := WSTRING#'';
   me.stations[27].raw[3,5] := WSTRING#'';
   me.stations[27].raw[3,6] := WSTRING#'';
   me.stations[27].raw[3,7] := WSTRING#'';
   me.stations[27].raw[4,0] := WSTRING#'16.32.112.553.010A';
   me.stations[27].raw[4,1] := WSTRING#'16.32.112.553.020A';
   me.stations[27].raw[4,2] := WSTRING#'16.32.112.553.300C';
   me.stations[27].raw[4,3] := WSTRING#'16.32.112.553.100D';
   me.stations[27].raw[4,4] := WSTRING#'';
   me.stations[27].raw[4,5] := WSTRING#'';
   me.stations[27].raw[4,6] := WSTRING#'';
   me.stations[27].raw[4,7] := WSTRING#'';
   me.stations[27].raw[5,0] := WSTRING#'16.32.112.553.220A';
   me.stations[27].raw[5,1] := WSTRING#'16.32.112.553.100D';
   me.stations[27].raw[5,2] := WSTRING#'16.32.112.054.041A';
   me.stations[27].raw[5,3] := WSTRING#'16.32.112.057.010A';
   me.stations[27].raw[5,4] := WSTRING#'';
   me.stations[27].raw[5,5] := WSTRING#'';
   me.stations[27].raw[5,6] := WSTRING#'';
   me.stations[27].raw[5,7] := WSTRING#'';
   me.stations[27].raw[6,0] := WSTRING#'16.32.112.553.220A';
   me.stations[27].raw[6,1] := WSTRING#'16.32.112.553.100D';
   me.stations[27].raw[6,2] := WSTRING#'16.32.112.054.041A';
   me.stations[27].raw[6,3] := WSTRING#'16.32.112.057.010A';
   me.stations[27].raw[6,4] := WSTRING#'';
   me.stations[27].raw[6,5] := WSTRING#'';
   me.stations[27].raw[6,6] := WSTRING#'';
   me.stations[27].raw[6,7] := WSTRING#'';
   me.stations[27].raw[7,0] := WSTRING#'16.32.112.503.220A';
   me.stations[27].raw[7,1] := WSTRING#'16.32.112.516.110E';
   me.stations[27].raw[7,2] := WSTRING#'16.32.112.536.010A';
   me.stations[27].raw[7,3] := WSTRING#'';
   me.stations[27].raw[7,4] := WSTRING#'';
   me.stations[27].raw[7,5] := WSTRING#'';
   me.stations[27].raw[7,6] := WSTRING#'';
   me.stations[27].raw[7,7] := WSTRING#'';
   me.stations[27].raw[8,0] := WSTRING#'16.32.112.503.210A';
   me.stations[27].raw[8,1] := WSTRING#'16.32.112.543.210E';
   me.stations[27].raw[8,2] := WSTRING#'16.32.112.543.020A';
   me.stations[27].raw[8,3] := WSTRING#'';
   me.stations[27].raw[8,4] := WSTRING#'';
   me.stations[27].raw[8,5] := WSTRING#'';
   me.stations[27].raw[8,6] := WSTRING#'';
   me.stations[28].raw[0,0] := WSTRING#'11.52.001.315.000B';
   me.stations[28].raw[0,1] := WSTRING#'11.52.001.316.001D';
   me.stations[28].raw[0,2] := WSTRING#'11.52.001.0545.000B';
   me.stations[28].raw[0,3] := WSTRING#'';
   me.stations[28].raw[0,4] := WSTRING#'';
   me.stations[28].raw[0,5] := WSTRING#'';
   me.stations[28].raw[0,6] := WSTRING#'';
   me.stations[28].raw[0,7] := WSTRING#'';
   me.stations[28].raw[1,0] := WSTRING#'11.54.017.315.001F';
   me.stations[28].raw[1,1] := WSTRING#'11.54.007.315.026G';
   me.stations[28].raw[1,2] := WSTRING#'11.54.007.045.015D';
   me.stations[28].raw[1,3] := WSTRING#'11.54.007.052.007B';
   me.stations[28].raw[1,4] := WSTRING#'11.54.007.052.008A';
   me.stations[28].raw[1,5] := WSTRING#'';
   me.stations[28].raw[1,6] := WSTRING#'';
   me.stations[28].raw[1,7] := WSTRING#'';
   me.stations[28].raw[2,0] := WSTRING#'11.54.017.315.001F';
   me.stations[28].raw[2,1] := WSTRING#'11.54.007.315.026G';
   me.stations[28].raw[2,2] := WSTRING#'11.54.007.045.015D';
   me.stations[28].raw[2,3] := WSTRING#'11.54.007.052.009B';
   me.stations[28].raw[2,4] := WSTRING#'11.54.007.052.010B';
   me.stations[28].raw[2,5] := WSTRING#'';
   me.stations[28].raw[2,6] := WSTRING#'';
   me.stations[28].raw[2,7] := WSTRING#'';
   // me.stations[0] : volvo 16 01
   // me.stations[1] : volvo 16 02
   // me.stations[2] : volvo 16 03
   // me.stations[3] : volvo 16 04
   // me.stations[4] : volvo 16 05
   // me.stations[5] : volvo 16 06
   // me.stations[6] : volvo 16 07
   // me.stations[7] : volvo 16 08
   // me.stations[8] : volvo 16 09
   // me.stations[9] : volvo 16 10
   // me.stations[10] : volvo 16 11
   // me.stations[11] : chm 01
   // me.stations[12] : chm 02
   // me.stations[13] : chm 03
   // me.stations[14] : chm 04
   // me.stations[15] : cdo 01
   // me.stations[16] : cdo 02
   // me.stations[17] : cdo 03
   // me.stations[18] : bfl 01
   // me.stations[19] : bfl 02
   // me.stations[20] : bfl 03
   // me.stations[21] : lgs 01
   // me.stations[22] : lgs 02
   // me.stations[23] : lgs 03
   // me.stations[24] : cv 01
   // me.stations[25] : cv 02
   // me.stations[26] : cv 03
   // me.stations[27] : cv 04
   // me.stations[28] : pc 01
   // me.stations[29] : pc 02
END_DATA_BLOCK

// folder: Network Diagnostics

DATA_BLOCK "Net Diag: Global"   // DB7
{ S7_Optimized_Access := 'TRUE' }
VERSION : 0.1
   VAR
      plcData : "UserDiag_typePLC";   // PLC diagnostics data
      ioSystemData : Array[1.."USERDIAG_IO_SYSTEMS_UPPER_LIM"] of "UserDiag_typeIOSystem";   // IO-System diagnostics data
      startDiag : Bool := false;   // Startflag for diagnostic
   END_VAR
BEGIN
END_DATA_BLOCK

DATA_BLOCK "Net Diag: Startup"   // DB8
{ S7_Optimized_Access := 'TRUE' }
VERSION : 0.1
// stored: InstanceOfName NetDiag: Coordinate
"NetDiag: Coordinate"
BEGIN
END_DATA_BLOCK

// folder: (top level)

FUNCTION_BLOCK "EMP"   // FB1, LAD
{ S7_Optimized_Access := 'TRUE' }
VERSION : 0.1
   VAR
      instAniPNTmr : "Animate: PN & Timers";
      instBaseAni : "Base Animations";
      instClrReqData : "Clear Part Requests";
      instClpseTable : "Collapse Table";
      instDfltTmrPrst : "Load Default Timer Presets";
      instHMIAni : "Format Part Call Requests";
      instHMIBarcode : "HMI Barcod Screen";
      instHMISettings : "HMI Settings Screen";
      instInitialize : "Initialize";
      instKP8BtnAct : "KP8 Button Activation";
      instKP8Drvs : Array[0.."stnCount"] of "KP8 Driver";
      instKP8ExpAni : "KP8 Expanded Animations";
      instPartTimers : "Part Timers";
      instPopulateHMI : "HMI Populate Part Call";
      instPopulateLED : "LED Populate Sign";
      instRcrdPartReq : "Record Part Request";
      instRmvPartReq : "Remove Part Request";
      instRstInitReq : "Reset Init Requests";
      instSLAni : "Stack Light Animations";
   END_VAR
   VAR RETAIN
      stations : "Stations";
   END_VAR
   VAR
      instGlblToSim : "Global to Sim";
      instLogReq : "Buffer Log: Part Requests";
      instUserDiag_Diag : "NetDiag: Coordinate";
      instUserDiagGetIPAddress : "NetDiag: Get IPs";
      statStartDiag : Bool := false;   // Static start Diagnostics
      instNetHealthScreen : "HMI: Network Health";
      instHMIStationDriver : "HSS: Driver";
   END_VAR
   VAR_TEMP
      i : Int;
   END_VAR
BEGIN

REGION Network 1: Static start Diagnostics
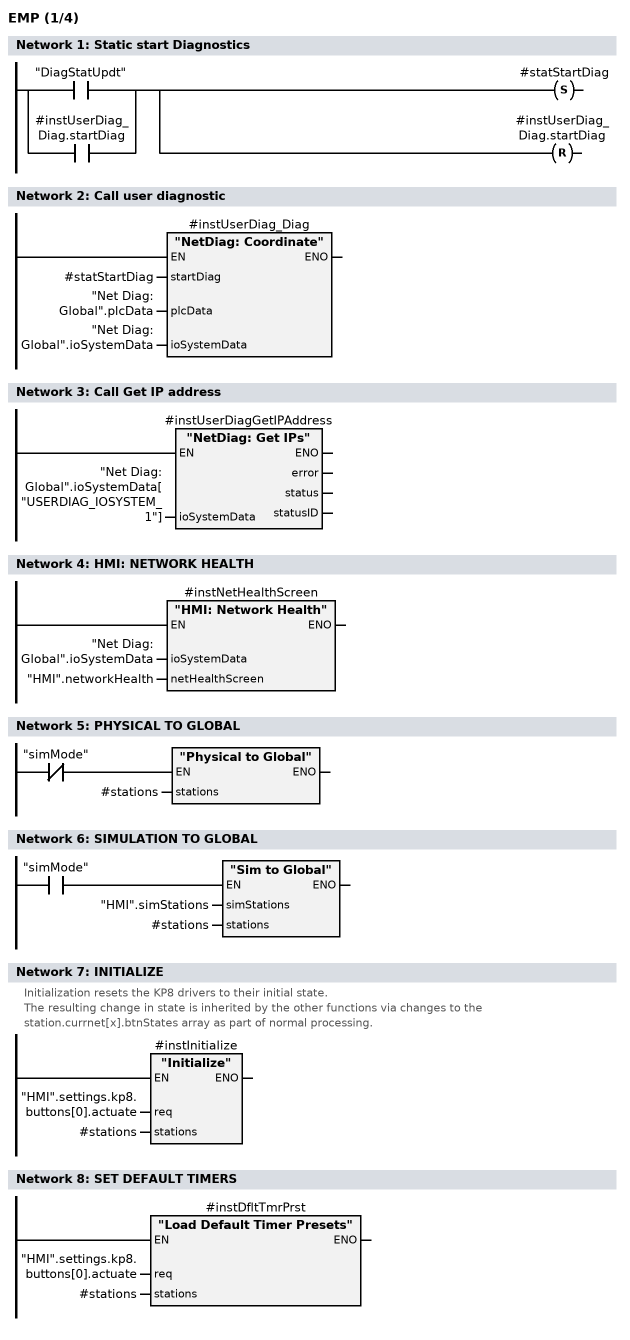
   RUNG wire#powerrail
      Contact( "DiagStatUpdt" )
      wire#w1
      S_Coil( #statStartDiag )
   END_RUNG
   RUNG wire#powerrail
      Contact( #instUserDiag_Diag.startDiag )
   END_RUNG wire#w1
   RUNG wire#w1
      R_Coil( #instUserDiag_Diag.startDiag )
   END_RUNG
   // the same network as SCL:
   IF "DiagStatUpdt" OR #instUserDiag_Diag.startDiag THEN
       #statStartDiag := TRUE;
       #instUserDiag_Diag.startDiag := FALSE;
   END_IF;
END_REGION

REGION Network 2: Call user diagnostic
   RUNG wire#powerrail
      #instUserDiag_Diag(startDiag := #statStartDiag, plcData := "Net Diag: Global".plcData, ioSystemData := "Net Diag: Global".ioSystemData)
   END_RUNG
   // the same network as SCL:
   #instUserDiag_Diag(startDiag := #statStartDiag,   // "NetDiag: Coordinate"
                      plcData := "Net Diag: Global".plcData,
                      ioSystemData := "Net Diag: Global".ioSystemData);
END_REGION

REGION Network 3: Call Get IP address
   RUNG wire#powerrail
      #instUserDiagGetIPAddress(ioSystemData := "Net Diag: Global".ioSystemData["USERDIAG_IOSYSTEM_1"], error =>, status =>, statusID =>)
   END_RUNG
   // the same network as SCL:
   #instUserDiagGetIPAddress(ioSystemData := "Net Diag: Global".ioSystemData["USERDIAG_IOSYSTEM_1"]);   // "NetDiag: Get IPs"
END_REGION

REGION Network 4: HMI: NETWORK HEALTH
   RUNG wire#powerrail
      #instNetHealthScreen(ioSystemData := "Net Diag: Global".ioSystemData, netHealthScreen := "HMI".networkHealth)
   END_RUNG
   // the same network as SCL:
   #instNetHealthScreen(ioSystemData := "Net Diag: Global".ioSystemData, netHealthScreen := "HMI".networkHealth);   // "HMI: Network Health"
END_REGION

REGION Network 5: PHYSICAL TO GLOBAL
   RUNG wire#powerrail
      I_Contact( "simMode" )
      "Physical to Global"(stations := #stations)
   END_RUNG
   // the same network as SCL:
   IF NOT "simMode" THEN "Physical to Global"(stations := #stations); END_IF;
END_REGION

REGION Network 6: SIMULATION TO GLOBAL
   RUNG wire#powerrail
      Contact( "simMode" )
      "Sim to Global"(simStations := "HMI".simStations, stations := #stations)
   END_RUNG
   // the same network as SCL:
   IF "simMode" THEN "Sim to Global"(simStations := "HMI".simStations, stations := #stations); END_IF;
END_REGION

REGION Network 7: INITIALIZE
   // Initialization resets the KP8 drivers to their initial state.
   // The resulting change in state is inherited by the other functions via changes to the
   // station.currnet[x].btnStates array as part of normal processing.
   RUNG wire#powerrail
      #instInitialize(req := "HMI".settings.kp8.buttons[0].actuate, stations := #stations)
   END_RUNG
   // the same network as SCL:
   #instInitialize(req := "HMI".settings.kp8.buttons[0].actuate, stations := #stations);   // "Initialize"
END_REGION

REGION Network 8: SET DEFAULT TIMERS
   RUNG wire#powerrail
      #instDfltTmrPrst(req := "HMI".settings.kp8.buttons[0].actuate, stations := #stations)
   END_RUNG
   // the same network as SCL:
   #instDfltTmrPrst(req := "HMI".settings.kp8.buttons[0].actuate, stations := #stations);   // "Load Default Timer Presets"
END_REGION

REGION Network 9: CLEAR PART REQUEST DATA